// TIA Portal project "proiect" (V17) (continued)
   // ASSB[18] := 18;
   // ASSB[19] := 19;
   // ASSB[20] := 20;
   // ASSB[21] := 21;
   // ASSB[22] := 22;
   // ASSB[23] := 23;
   // ASSB[24] := 24;
   // ASSB[25] := 25;
   // ASSB[26] := 26;
   // ASSB[27] := 27;
   // ASSB[28] := 28;
   // ASSB[29] := 29;
   // ASSB[30] := 30;
   // ASSB[31] := 31;
   // ASSB[32] := 32;
   // ASSB[33] := 33;
   // ASSB[34] := 34;
   // ASSB[35] := 35;
   // ASSB[36] := 36;
   // ASSB[37] := 37;
   // ASSB[38] := 38;
   // ASSB[39] := 39;
   // ASSB[40] := 40;
   // ASSB[41] := 41;
   // ASSB[42] := 42;
   // ASSB[43] := 43;
   // ASSB[44] := 44;
   // ASSB[45] := 45;
   // ASSB[46] := 46;
   // ASSB[47] := 47;
   // ASSB[48] := 48;
   // ASSB[49] := 49;
   // ASSB[50] := 50;
   // ASSB[51] := 51;
   // ASSB[52] := 52;
   // ASSB[53] := 53;
   // ASSB[54] := 54;
   // ASSB[55] := 55;
   // ASSB[56] := 56;
   // ASSB[57] := 57;
   // ASSB[58] := 58;
   // ASSB[59] := 59;
   // ASSB[60] := 60;
   // ASSB[61] := 61;
   // ASSB[62] := 62;
   // ASSB[63] := 63;
   // ASSB[64] := 64;
   // ASSB[65] := 65;
   // ASSB[66] := 66;
   // ASSB[67] := 67;
   // ASSB[68] := 68;
   // ASSB[69] := 69;
   // ASSB[70] := 70;
   // ASSB[71] := 71;
   // ASSB[72] := 72;
   // ASSB[73] := 73;
   // ASSB[74] := 74;
   // ASSB[75] := 75;
   // ASSB[76] := 76;
   // ASSB[77] := 77;
   // PTTS[5] := 2;
   // PTTS[6] := 3;
   // PTTS[7] := 4;
   // PTTS[8] := 5;
   // PTTS[9] := 6;
   // PTTS[10] := 7;
   // PTTS[11] := 72;
   // PTTS[12] := 9;
   // PTTS[13] := 10;
   // PTTS[14] := 11;
   // PTTS[15] := 98;
   // PTTS[16] := 13;
   // PTTS[17] := 14;
   // PTTS[18] := 15;
   // PTTS[19] := 16;
   // PTTS[20] := 17;
   // PTTS[21] := 19;
   // PTTS[22] := 20;
   // PTTS[23] := 21;
   // PTTS[24] := 22;
   // PTTS[25] := 23;
   // PTTS[26] := 24;
   // PTTS[27] := 69;
   // PTTS[28] := 26;
   // PTTS[29] := 27;
   // PTTS[30] := 28;
   // PTTS[31] := 97;
   // PTTS[32] := 30;
   // PTTS[33] := 31;
   // PTTS[34] := 32;
   // PTTS[35] := 33;
   // PTTS[36] := 34;
   // PTTS[37] := 36;
   // PTTS[38] := 37;
   // PTTS[39] := 38;
   // PTTS[40] := 68;
   // PTTS[41] := 40;
   // PTTS[42] := 41;
   // PTTS[43] := 42;
   // PTTS[44] := 96;
   // PTTS[45] := 44;
   // PTTS[46] := 45;
   // PTTS[47] := 46;
   // PTTS[48] := 47;
   // PTTS[49] := 48;
   // PTTS[50] := 53;
   // PTTS[51] := 55;
   // PTTS[52] := 99;
   // PTTS[53] := 57;
   // PTTS[54] := 58;
   // PTTS[55] := 54;
   // PTTS[56] := 59;
   // PTTS[57] := 60;
   // PTTS[58] := 255;
   // PTTS[59] := 62;
   // PTTS[60] := 39;
   // PTTS[61] := 64;
   // PTTS[62] := 66;
   // PTTS[63] := 67;
   // PTTS[64] := 8;
   // PTTS[65] := 25;
   // PTTS[66] := 70;
   // PTTS[67] := 71;
   // PTTS[68] := 73;
   // PTTS[69] := 74;
   // PTTS[70] := 1;
   // PTTS[71] := 63;
   // PTTS[72] := 76;
   // PTTS[73] := 78;
   // PTTS[74] := 43;
   // PTTS[75] := 49;
   // PTTS[76] := 80;
   // PTTS[77] := 29;
   // NTTS[5] := 3;
   // NTTS[6] := 4;
   // NTTS[7] := 5;
   // NTTS[8] := 6;
   // NTTS[9] := 7;
   // NTTS[10] := 8;
   // NTTS[11] := 9;
   // NTTS[12] := 10;
   // NTTS[13] := 11;
   // NTTS[14] := 12;
   // NTTS[15] := 13;
   // NTTS[16] := 14;
   // NTTS[17] := 15;
   // NTTS[18] := 16;
   // NTTS[19] := 17;
   // NTTS[20] := 18;
   // NTTS[21] := 20;
   // NTTS[22] := 21;
   // NTTS[23] := 22;
   // NTTS[24] := 23;
   // NTTS[25] := 24;
   // NTTS[26] := 25;
   // NTTS[27] := 26;
   // NTTS[28] := 27;
   // NTTS[29] := 28;
   // NTTS[30] := 29;
   // NTTS[31] := 30;
   // NTTS[32] := 31;
   // NTTS[33] := 32;
   // NTTS[34] := 33;
   // NTTS[35] := 34;
   // NTTS[36] := 35;
   // NTTS[37] := 37;
   // NTTS[38] := 38;
   // NTTS[39] := 39;
   // NTTS[40] := 40;
   // NTTS[41] := 41;
   // NTTS[42] := 42;
   // NTTS[43] := 78;
   // NTTS[44] := 44;
   // NTTS[45] := 45;
   // NTTS[46] := 46;
   // NTTS[47] := 47;
   // NTTS[48] := 48;
   // NTTS[49] := 49;
   // NTTS[50] := 55;
   // NTTS[51] := 56;
   // NTTS[52] := 57;
   // NTTS[53] := 58;
   // NTTS[54] := 54;
   // NTTS[55] := 59;
   // NTTS[56] := 60;
   // NTTS[57] := 61;
   // NTTS[58] := 62;
   // NTTS[59] := 63;
   // NTTS[60] := 66;
   // NTTS[61] := 65;
   // NTTS[62] := 67;
   // NTTS[63] := 68;
   // NTTS[64] := 73;
   // NTTS[65] := 70;
   // NTTS[66] := 71;
   // NTTS[67] := 69;
   // NTTS[68] := 74;
   // NTTS[69] := 72;
   // NTTS[70] := 36;
   // NTTS[71] := 76;
   // NTTS[72] := 77;
   // NTTS[73] := 43;
   // NTTS[74] := 79;
   // NTTS[75] := 80;
   // NTTS[76] := 81;
   // NTTS[77] := 82;
   // SW_SQTS[3] := 2;
   // SW_SQTS[4] := 2;
   // SW_SQTS[5] := 3;
   // SW_SQTS[6] := 3;
   // SW_SQTS[7] := 3;
   // SW_SQTS[8] := 3;
   // SW_SQTS[9] := 3;
   // SW_SQTS[10] := 3;
   // SW_SQTS[11] := 3;
   // SW_SQTS[12] := 3;
   // SW_SQTS[13] := 3;
   // SW_SQTS[14] := 3;
   // SW_SQTS[15] := 3;
   // SW_SQTS[16] := 3;
   // SW_SQTS[17] := 3;
   // SW_SQTS[18] := 3;
   // SW_SQTS[19] := 3;
   // SW_SQTS[20] := 3;
   // SW_SQTS[21] := 4;
   // SW_SQTS[22] := 4;
   // SW_SQTS[23] := 4;
   // SW_SQTS[24] := 4;
   // SW_SQTS[25] := 4;
   // SW_SQTS[26] := 4;
   // SW_SQTS[27] := 4;
   // SW_SQTS[28] := 4;
   // SW_SQTS[29] := 4;
   // SW_SQTS[30] := 4;
   // SW_SQTS[31] := 4;
   // SW_SQTS[32] := 4;
   // SW_SQTS[33] := 4;
   // SW_SQTS[34] := 4;
   // SW_SQTS[35] := 4;
   // SW_SQTS[36] := 4;
   // SW_SQTS[37] := 5;
   // SW_SQTS[38] := 5;
   // SW_SQTS[39] := 5;
   // SW_SQTS[40] := 5;
   // SW_SQTS[41] := 5;
   // SW_SQTS[42] := 5;
   // SW_SQTS[43] := 5;
   // SW_SQTS[44] := 5;
   // SW_SQTS[45] := 5;
   // SW_SQTS[46] := 5;
   // SW_SQTS[47] := 5;
   // SW_SQTS[48] := 5;
   // SW_SQTS[49] := 5;
   // SW_SQTS[50] := 2;
   // SW_SQTS[51] := 2;
   // SW_SQTS[52] := 2;
   // SW_SQTS[53] := 2;
   // SW_SQTS[54] := 2;
   // SW_SQTS[55] := 2;
   // SW_SQTS[56] := 2;
   // SW_SQTS[57] := 2;
   // SW_SQTS[58] := 6;
   // SW_SQTS[59] := 7;
   // SW_SQTS[60] := 5;
   // SW_SQTS[61] := 8;
   // SW_SQTS[62] := 5;
   // SW_SQTS[63] := 5;
   // SW_SQTS[64] := 3;
   // SW_SQTS[65] := 4;
   // SW_SQTS[66] := 4;
   // SW_SQTS[67] := 4;
   // SW_SQTS[68] := 3;
   // SW_SQTS[69] := 3;
   // SW_SQTS[70] := 9;
   // SW_SQTS[71] := 7;
   // SW_SQTS[72] := 7;
   // SW_SQTS[73] := 5;
   // SW_SQTS[74] := 5;
   // SW_SQTS[75] := 5;
   // SW_SQTS[76] := 5;
   // SW_SQTS[77] := 4;
   // SINI[2] := 255;
   // LSTT[83] := 255;
   // LSTT[84] := 255;
   // LSTT[86] := 255;
   // ATAJ[82] := 82;
   // ATAJ[83] := 83;
   // ATAJ[84] := 84;
   // ATAJ[85] := 85;
   // ATAJ[86] := 86;
   // ATAB[82] := 82;
   // ATAB[83] := 83;
   // ATAB[84] := 84;
   // ATAB[85] := 85;
   // ATAB[86] := 86;
   // PSTT[82] := 77;
   // PSTT[83] := 78;
   // PSTT[84] := 79;
   // PSTT[85] := 80;
   // PSTT[86] := 81;
   // NSTT[83] := 91;
   // NSTT[84] := 80;
   // NSTT[86] := 82;
   // ASSJ[78] := 78;
   // ASSJ[79] := 79;
   // ASSJ[80] := 80;
   // ASSJ[81] := 81;
   // ASSB[78] := 78;
   // ASSB[79] := 79;
   // ASSB[80] := 80;
   // ASSB[81] := 81;
   // PTTS[78] := 82;
   // PTTS[79] := 35;
   // PTTS[80] := 84;
   // PTTS[81] := 12;
   // NTTS[78] := 83;
   // NTTS[79] := 84;
   // NTTS[80] := 85;
   // NTTS[81] := 86;
   // SW_SQTS[78] := 4;
   // SW_SQTS[79] := 4;
   // SW_SQTS[80] := 4;
   // SW_SQTS[81] := 3;
   // SWITCH[0] := 192;
   // SWITCH[1] := 1;
   // SWITCH[2] := 14;
   // SWITCH[3] := 112;
   // SWITCH[4] := 128;
   // SWITCH[5] := 3;
   // SWITCH[6] := 28;
   // SWITCH[7] := 224;
   // LSTT[87] := 255;
   // LSTT[88] := 255;
   // LSTT[90] := 255;
   // LSTT[91] := 255;
   // LSTT[92] := 255;
   // LSTT[94] := 255;
   // ATAJ[87] := 87;
   // ATAJ[88] := 88;
   // ATAJ[89] := 89;
   // ATAJ[90] := 90;
   // ATAJ[91] := 91;
   // ATAJ[92] := 92;
   // ATAJ[93] := 93;
   // ATAJ[94] := 94;
   // ATAJ[95] := 95;
   // ATAB[87] := 87;
   // ATAB[88] := 88;
   // ATAB[89] := 89;
   // ATAB[90] := 90;
   // ATAB[91] := 91;
   // ATAB[92] := 92;
   // ATAB[93] := 93;
   // ATAB[95] := 95;
   // PSTT[87] := 82;
   // PSTT[88] := 83;
   // PSTT[89] := 84;
   // PSTT[90] := 85;
   // PSTT[91] := 86;
   // PSTT[92] := 87;
   // PSTT[93] := 88;
   // PSTT[95] := 89;
   // NSTT[87] := 92;
   // NSTT[88] := 84;
   // NSTT[90] := 86;
   // NSTT[91] := 93;
   // NSTT[92] := 88;
   // NSTT[94] := 89;
   // ASSJ[82] := 82;
   // ASSJ[83] := 83;
   // ASSJ[84] := 84;
   // ASSJ[85] := 85;
   // ASSJ[86] := 86;
   // ASSJ[87] := 87;
   // ASSJ[88] := 88;
   // ASSJ[89] := 89;
   // ASSB[82] := 82;
   // ASSB[83] := 83;
   // ASSB[84] := 84;
   // ASSB[85] := 85;
   // ASSB[86] := 86;
   // ASSB[87] := 87;
   // ASSB[88] := 88;
   // ASSB[89] := 89;
   // PTTS[82] := 86;
   // PTTS[83] := 18;
   // PTTS[84] := 88;
   // PTTS[85] := 56;
   // PTTS[86] := 90;
   // PTTS[87] := 61;
   // PTTS[88] := 92;
   // PTTS[89] := 94;
   // NTTS[82] := 87;
   // NTTS[83] := 88;
   // NTTS[84] := 89;
   // NTTS[85] := 90;
   // NTTS[86] := 91;
   // NTTS[87] := 92;
   // NTTS[88] := 93;
   // NTTS[89] := 95;
   // SW_SQTS[82] := 3;
   // SW_SQTS[83] := 3;
   // SW_SQTS[84] := 3;
   // SW_SQTS[85] := 2;
   // SW_SQTS[86] := 2;
   // SW_SQTS[87] := 2;
   // SW_SQTS[88] := 2;
   // SW_SQTS[89] := 10;
   // SW_SQTS[2] := 2;
   // SWITCH[8] := 252;
   // SWITCH[9] := 248;
   // SWITCH[10] := 199;
   // SW_SQTS[1] := 1;
   // ATAB[0] := 94;
   // SWITCH[12] := 6;
   // LSTT[61] := 255;
   // LSTT[43] := 255;
   // LSTT[22] := 255;
   // SWITCH[11] := 63;
   // NSTT[61] := 87;
   // NSTT[43] := 74;
   // NSTT[22] := 24;
   // SWITCH[13] := 14;
   // SWITCH[14] := 112;
   // LSTT[96] := 255;
   // LSTT[97] := 255;
   // LSTT[98] := 255;
   // LSTT[99] := 255;
   // ATAJ[96] := 96;
   // ATAJ[97] := 97;
   // ATAJ[98] := 98;
   // ATAJ[99] := 99;
   // ATAB[96] := 96;
   // ATAB[97] := 97;
   // ATAB[98] := 98;
   // ATAB[99] := 99;
   // PSTT[96] := 90;
   // PSTT[97] := 91;
   // PSTT[98] := 92;
   // PSTT[99] := 93;
   // NSTT[96] := 44;
   // NSTT[97] := 31;
   // NSTT[98] := 15;
   // NSTT[99] := 52;
   // ASSJ[90] := 90;
   // ASSJ[91] := 91;
   // ASSJ[92] := 92;
   // ASSJ[93] := 93;
   // ASSB[90] := 90;
   // ASSB[91] := 91;
   // ASSB[92] := 92;
   // ASSB[93] := 93;
   // PTTS[90] := 79;
   // PTTS[91] := 83;
   // PTTS[92] := 87;
   // PTTS[93] := 91;
   // NTTS[90] := 96;
   // NTTS[91] := 97;
   // NTTS[92] := 98;
   // NTTS[93] := 99;
   // SW_SQTS[90] := 5;
   // SW_SQTS[91] := 4;
   // SW_SQTS[92] := 3;
   // SW_SQTS[93] := 2;
BEGIN
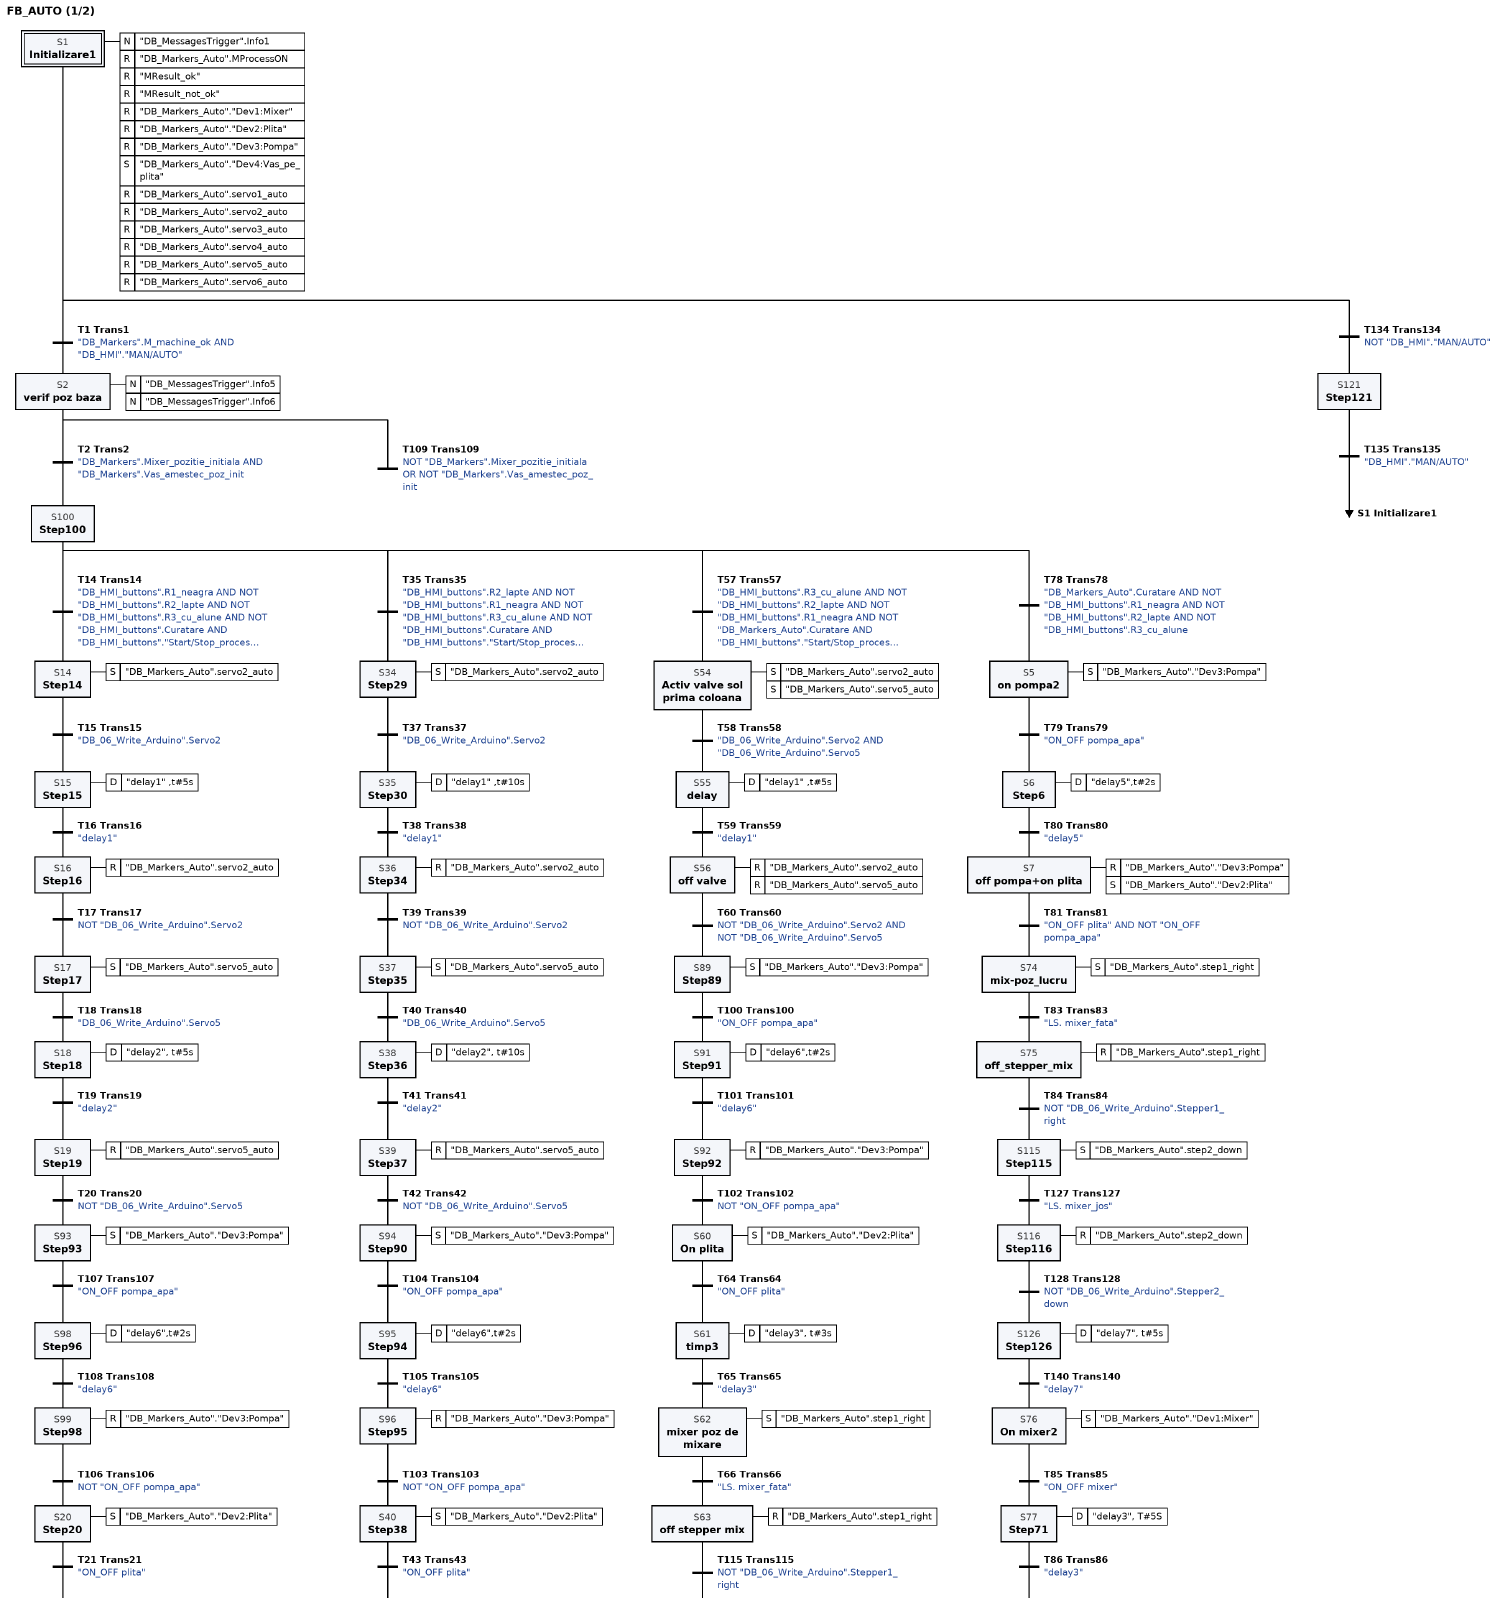
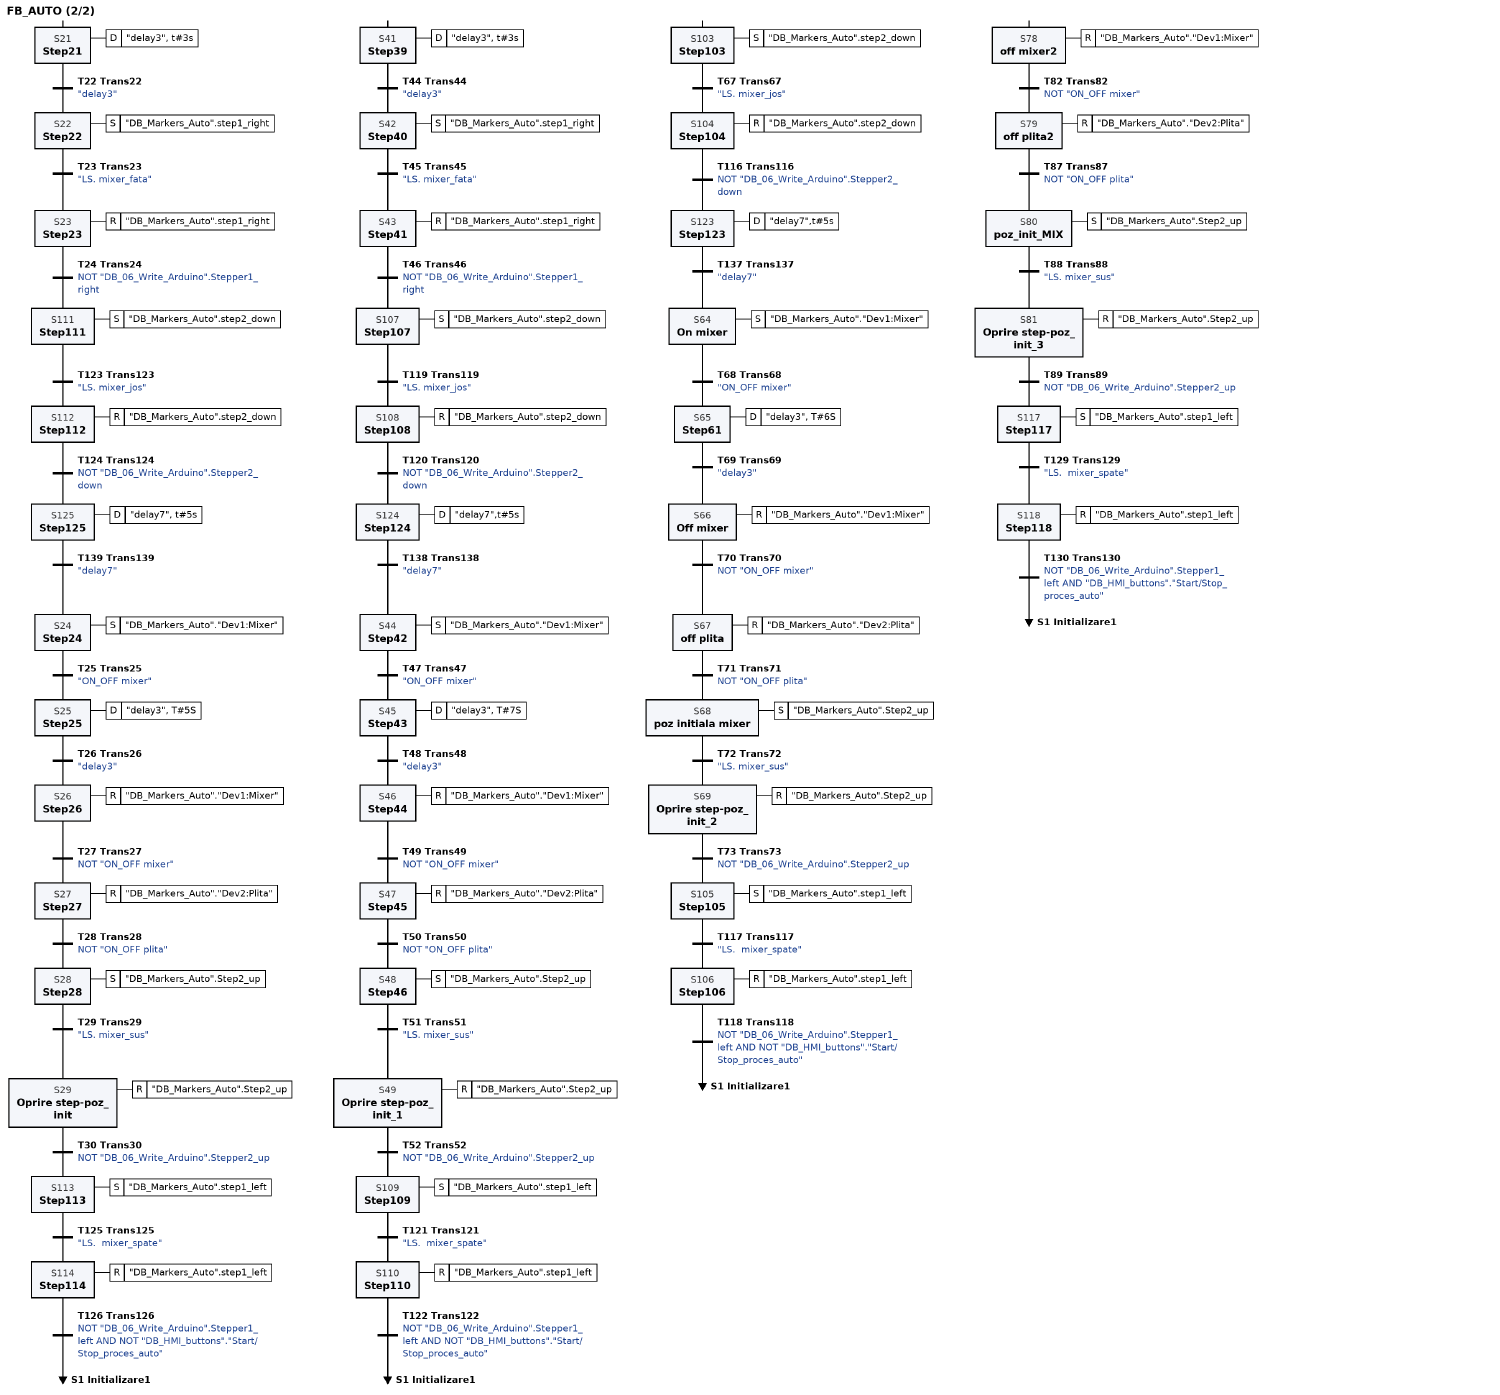
   // sequencer 1
   INITIAL_STEP Initializare1:   // S1, max time T#10S, warning time T#7S
      // Initializare
              N    "DB_MessagesTrigger".Info1
              R    "DB_Markers_Auto".MProcessON
              R    "MResult_ok"
              R    "MResult_not_ok"
              R    "DB_Markers_Auto"."Dev1:Mixer"
              R    "DB_Markers_Auto"."Dev2:Plita"
              R    "DB_Markers_Auto"."Dev3:Pompa"
              S    "DB_Markers_Auto"."Dev4:Vas_pe_plita"
              R    "DB_Markers_Auto".servo1_auto
              R    "DB_Markers_Auto".servo2_auto
              R    "DB_Markers_Auto".servo3_auto
              R    "DB_Markers_Auto".servo4_auto
              R    "DB_Markers_Auto".servo5_auto
              R    "DB_Markers_Auto".servo6_auto
              R    "DB_Markers_Auto".step1_left
              R    "DB_Markers_Auto".step1_right
              R    "DB_Markers_Auto".Step2_up
              R    "DB_Markers_Auto".step2_down
   END_STEP
   TRANSITION Trans1 FROM Initializare1 TO "verif poz baza"   // T1
      := "DB_Markers".M_machine_ok AND "DB_HMI"."MAN/AUTO";
   END_TRANSITION
   TRANSITION Trans134 FROM Initializare1 TO Step121   // T134
      := NOT "DB_HMI"."MAN/AUTO";
   END_TRANSITION
   STEP "verif poz baza":   // S2, max time T#10S, warning time T#7S
      // Verificare dispozitive in pozitia de baza
              N    "DB_MessagesTrigger".Info5
              N    "DB_MessagesTrigger".Info6
   END_STEP
   TRANSITION Trans2 FROM "verif poz baza" TO Step100   // T2
      := "DB_Markers".Mixer_pozitie_initiala AND "DB_Markers".Vas_amestec_poz_init;
   END_TRANSITION
   TRANSITION Trans109 FROM "verif poz baza" TO ?   // T109
      := NOT "DB_Markers".Mixer_pozitie_initiala OR NOT "DB_Markers".Vas_amestec_poz_init;
   END_TRANSITION
   STEP Step103:   // S103, max time T#10S, warning time T#7S
              S    "DB_Markers_Auto".step2_down
   END_STEP
   TRANSITION Trans67 FROM Step103 TO Step104   // T67
      := "LS. mixer_jos";
   END_TRANSITION
   STEP Step29:   // S34, max time T#10S, warning time T#7S
      // Activare valve solutii rand superior
              S    "DB_Markers_Auto".servo2_auto
   END_STEP
   TRANSITION Trans37 FROM Step29 TO Step30   // T37
      := "DB_06_Write_Arduino".Servo2;
   END_TRANSITION
   STEP Step14:   // S14, max time T#10S, warning time T#7S
      // Activare valve solutii rand superior
              S    "DB_Markers_Auto".servo2_auto
   END_STEP
   TRANSITION Trans15 FROM Step14 TO Step15   // T15
      := "DB_06_Write_Arduino".Servo2;
   END_TRANSITION
   STEP Step15:   // S15, max time T#10S, warning time T#7S
      // delay
              D    "delay1" ,t#5s
   END_STEP
   TRANSITION Trans16 FROM Step15 TO Step16   // T16
      := "delay1";
   END_TRANSITION
   STEP Step16:   // S16, max time T#10S, warning time T#7S
      // inchidere valve rand superior
              R    "DB_Markers_Auto".servo2_auto
   END_STEP
   TRANSITION Trans17 FROM Step16 TO Step17   // T17
      := NOT "DB_06_Write_Arduino".Servo2;
   END_TRANSITION
   STEP Step17:   // S17, max time T#10S, warning time T#7S
      // deschidere valve solutii rand inferior
              S    "DB_Markers_Auto".servo5_auto
   END_STEP
   TRANSITION Trans18 FROM Step17 TO Step18   // T18
      := "DB_06_Write_Arduino".Servo5;
   END_TRANSITION
   STEP Step18:   // S18, max time T#10S, warning time T#7S
      // delay
              D    "delay2", t#5s
   END_STEP
   TRANSITION Trans19 FROM Step18 TO Step19   // T19
      := "delay2";
   END_TRANSITION
   STEP Step19:   // S19, max time T#10S, warning time T#7S
      // inchidere valve rand inferior
              R    "DB_Markers_Auto".servo5_auto
   END_STEP
   TRANSITION Trans20 FROM Step19 TO Step93   // T20
      := NOT "DB_06_Write_Arduino".Servo5;
   END_TRANSITION
   STEP Step20:   // S20, max time T#10S, warning time T#7S
      // deschidere plita
              S    "DB_Markers_Auto"."Dev2:Plita"
   END_STEP
   TRANSITION Trans21 FROM Step20 TO Step21   // T21
      := "ON_OFF plita";
   END_TRANSITION
   STEP Step21:   // S21, max time T#10S, warning time T#7S
      // delay
              D    "delay3", t#3s
   END_STEP
   TRANSITION Trans22 FROM Step21 TO Step22   // T22
      := "delay3";
   END_TRANSITION
   STEP Step22:   // S22, max time T#10S, warning time T#7S
      // pozitionare mixer/pornire stepper
              S    "DB_Markers_Auto".step1_right
   END_STEP
   TRANSITION Trans23 FROM Step22 TO Step23   // T23
      := "LS. mixer_fata";
   END_TRANSITION
   STEP Step23:   // S23, max time T#10S, warning time T#7S
      // Oprire stepper/mixer
              R    "DB_Markers_Auto".step1_right
   END_STEP
   TRANSITION Trans24 FROM Step23 TO Step111   // T24
      := NOT "DB_06_Write_Arduino".Stepper1_right;
   END_TRANSITION
   STEP Step24:   // S24, max time T#10S, warning time T#7S
      // Pornire mixer(on,off)
              S    "DB_Markers_Auto"."Dev1:Mixer"
   END_STEP
   TRANSITION Trans25 FROM Step24 TO Step25   // T25
      := "ON_OFF mixer";
   END_TRANSITION
   STEP Step25:   // S25, max time T#10S, warning time T#7S
      // Delay(timp de mixare)
              D    "delay3", T#5S
   END_STEP
   TRANSITION Trans26 FROM Step25 TO Step26   // T26
      := "delay3";
   END_TRANSITION
   STEP Step26:   // S26, max time T#10S, warning time T#7S
      // Oprire mixer
              R    "DB_Markers_Auto"."Dev1:Mixer"
   END_STEP
   TRANSITION Trans27 FROM Step26 TO Step27   // T27
      := NOT "ON_OFF mixer";
   END_TRANSITION
   STEP Step27:   // S27, max time T#10S, warning time T#7S
      // Oprire plita
              R    "DB_Markers_Auto"."Dev2:Plita"
   END_STEP
   TRANSITION Trans28 FROM Step27 TO Step28   // T28
      := NOT "ON_OFF plita";
   END_TRANSITION
   STEP Step28:   // S28, max time T#10S, warning time T#7S
      // RETRAGERE MIXER IN POZITIA INITIALA
              S    "DB_Markers_Auto".Step2_up
   END_STEP
   TRANSITION Trans29 FROM Step28 TO "Oprire step-poz_init"   // T29
      := "LS. mixer_sus";
   END_TRANSITION
   STEP "Oprire step-poz_init":   // S29, max time T#10S, warning time T#7S
      // Oprire Stepper_pozitie initiala
              R    "DB_Markers_Auto".Step2_up
   END_STEP
   TRANSITION Trans30 FROM "Oprire step-poz_init" TO Step113   // T30
      := NOT "DB_06_Write_Arduino".Stepper2_up;
   END_TRANSITION
   STEP Step30:   // S35, max time T#10S, warning time T#7S
      // delay
              D    "delay1" ,t#10s
   END_STEP
   TRANSITION Trans38 FROM Step30 TO Step34   // T38
      := "delay1";
   END_TRANSITION
   STEP Step34:   // S36, max time T#10S, warning time T#7S
      // inchidere valve rand superior
              R    "DB_Markers_Auto".servo2_auto
   END_STEP
   TRANSITION Trans39 FROM Step34 TO Step35   // T39
      := NOT "DB_06_Write_Arduino".Servo2;
   END_TRANSITION
   STEP Step35:   // S37, max time T#10S, warning time T#7S
      // deschidere valve solutii rand inferior
              S    "DB_Markers_Auto".servo5_auto
   END_STEP
   TRANSITION Trans40 FROM Step35 TO Step36   // T40
      := "DB_06_Write_Arduino".Servo5;
   END_TRANSITION
   STEP Step36:   // S38, max time T#10S, warning time T#7S
      // delay
              D    "delay2", t#10s
   END_STEP
   TRANSITION Trans41 FROM Step36 TO Step37   // T41
      := "delay2";
   END_TRANSITION
   STEP Step37:   // S39, max time T#10S, warning time T#7S
      // inchidere valve rand inferior
              R    "DB_Markers_Auto".servo5_auto
   END_STEP
   TRANSITION Trans42 FROM Step37 TO Step90   // T42
      := NOT "DB_06_Write_Arduino".Servo5;
   END_TRANSITION
   STEP Step38:   // S40, max time T#10S, warning time T#7S
      // deschidere plita
              S    "DB_Markers_Auto"."Dev2:Plita"
   END_STEP
   TRANSITION Trans43 FROM Step38 TO Step39   // T43
      := "ON_OFF plita";
   END_TRANSITION
   STEP Step39:   // S41, max time T#10S, warning time T#7S
      // delay
              D    "delay3", t#3s
   END_STEP
   TRANSITION Trans44 FROM Step39 TO Step40   // T44
      := "delay3";
   END_TRANSITION
   STEP Step40:   // S42, max time T#10S, warning time T#7S
      // pozitionare mixer/pornire stepper
              S    "DB_Markers_Auto".step1_right
   END_STEP
   TRANSITION Trans45 FROM Step40 TO Step41   // T45
      := "LS. mixer_fata";
   END_TRANSITION
   STEP Step41:   // S43, max time T#10S, warning time T#7S
      // Oprire stepper/mixer
              R    "DB_Markers_Auto".step1_right
   END_STEP
   TRANSITION Trans46 FROM Step41 TO Step107   // T46
      := NOT "DB_06_Write_Arduino".Stepper1_right;
   END_TRANSITION
   STEP Step42:   // S44, max time T#10S, warning time T#7S
      // Pornire mixer(on,off)
              S    "DB_Markers_Auto"."Dev1:Mixer"
   END_STEP
   TRANSITION Trans47 FROM Step42 TO Step43   // T47
      := "ON_OFF mixer";
   END_TRANSITION
   STEP Step43:   // S45, max time T#10S, warning time T#7S
      // Delay(timp de mixare)
              D    "delay3", T#7S
   END_STEP
   TRANSITION Trans48 FROM Step43 TO Step44   // T48
      := "delay3";
   END_TRANSITION
   STEP Step44:   // S46, max time T#10S, warning time T#7S
      // Oprire mixer
              R    "DB_Markers_Auto"."Dev1:Mixer"
   END_STEP
   TRANSITION Trans49 FROM Step44 TO Step45   // T49
      := NOT "ON_OFF mixer";
   END_TRANSITION
   STEP Step45:   // S47, max time T#10S, warning time T#7S
      // Oprire plita
              R    "DB_Markers_Auto"."Dev2:Plita"
   END_STEP
   TRANSITION Trans50 FROM Step45 TO Step46   // T50
      := NOT "ON_OFF plita";
   END_TRANSITION
   STEP Step46:   // S48, max time T#10S, warning time T#7S
      // RETRAGERE MIXER IN POZITIA INITIALA
              S    "DB_Markers_Auto".Step2_up
   END_STEP
   TRANSITION Trans51 FROM Step46 TO "Oprire step-poz_init_1"   // T51
      := "LS. mixer_sus";
   END_TRANSITION
   STEP "Oprire step-poz_init_1":   // S49, max time T#10S, warning time T#7S
      // Oprire Stepper_pozitie initiala
              R    "DB_Markers_Auto".Step2_up
   END_STEP
   TRANSITION Trans52 FROM "Oprire step-poz_init_1" TO Step109   // T52
      := NOT "DB_06_Write_Arduino".Stepper2_up;
   END_TRANSITION
   STEP "Activ valve sol prima coloana":   // S54, max time T#10S, warning time T#7S
      // Activare valve solutii prima coloana
              S    "DB_Markers_Auto".servo2_auto
              S    "DB_Markers_Auto".servo5_auto
   END_STEP
   TRANSITION Trans58 FROM "Activ valve sol prima coloana" TO delay   // T58
      := "DB_06_Write_Arduino".Servo2 AND "DB_06_Write_Arduino".Servo5;
   END_TRANSITION
   STEP delay:   // S55, max time T#10S, warning time T#7S
      // delay
              D    "delay1" ,t#5s
   END_STEP
   TRANSITION Trans59 FROM delay TO "off valve"   // T59
      := "delay1";
   END_TRANSITION
   STEP "off valve":   // S56, max time T#10S, warning time T#7S
      // inchidere valve coloana 1
              R    "DB_Markers_Auto".servo2_auto
              R    "DB_Markers_Auto".servo5_auto
   END_STEP
   TRANSITION Trans60 FROM "off valve" TO Step89   // T60
      := NOT "DB_06_Write_Arduino".Servo2 AND NOT "DB_06_Write_Arduino".Servo5;
   END_TRANSITION
   STEP "On plita":   // S60, max time T#10S, warning time T#7S
      // deschidere plita
              S    "DB_Markers_Auto"."Dev2:Plita"
   END_STEP
   TRANSITION Trans64 FROM "On plita" TO timp3   // T64
      := "ON_OFF plita";
   END_TRANSITION
   STEP timp3:   // S61, max time T#10S, warning time T#7S
      // delay
              D    "delay3", t#3s
   END_STEP
   TRANSITION Trans65 FROM timp3 TO "mixer poz de mixare"   // T65
      := "delay3";
   END_TRANSITION
   STEP "mixer poz de mixare":   // S62, max time T#10S, warning time T#7S
      // pozitionare mixer/pornire stepper
              S    "DB_Markers_Auto".step1_right
   END_STEP
   TRANSITION Trans66 FROM "mixer poz de mixare" TO "off stepper mix"   // T66
      := "LS. mixer_fata";
   END_TRANSITION
   STEP "off stepper mix":   // S63, max time T#10S, warning time T#7S
      // Oprire stepper/mixer
              R    "DB_Markers_Auto".step1_right
   END_STEP
   TRANSITION Trans115 FROM "off stepper mix" TO Step103   // T115
      := NOT "DB_06_Write_Arduino".Stepper1_right;
   END_TRANSITION
   STEP "On mixer":   // S64, max time T#10S, warning time T#7S
      // Pornire mixer(on,off)
              S    "DB_Markers_Auto"."Dev1:Mixer"
   END_STEP
   TRANSITION Trans68 FROM "On mixer" TO Step61   // T68
      := "ON_OFF mixer";
   END_TRANSITION
   STEP Step61:   // S65, max time T#10S, warning time T#7S
      // Delay(timp de mixare)
              D    "delay3", T#6S
   END_STEP
   TRANSITION Trans69 FROM Step61 TO "Off mixer"   // T69
      := "delay3";
   END_TRANSITION
   STEP "Off mixer":   // S66, max time T#10S, warning time T#7S
      // Oprire mixer
              R    "DB_Markers_Auto"."Dev1:Mixer"
   END_STEP
   TRANSITION Trans70 FROM "Off mixer" TO "off plita"   // T70
      := NOT "ON_OFF mixer";
   END_TRANSITION
   STEP "off plita":   // S67, max time T#10S, warning time T#7S
      // Oprire plita
              R    "DB_Markers_Auto"."Dev2:Plita"
   END_STEP
   TRANSITION Trans71 FROM "off plita" TO "poz initiala mixer"   // T71
      := NOT "ON_OFF plita";
   END_TRANSITION
   STEP "poz initiala mixer":   // S68, max time T#10S, warning time T#7S
      // RETRAGERE MIXER IN POZITIA INITIALA
              S    "DB_Markers_Auto".Step2_up
   END_STEP
   TRANSITION Trans72 FROM "poz initiala mixer" TO "Oprire step-poz_init_2"   // T72
      := "LS. mixer_sus";
   END_TRANSITION
   STEP "Oprire step-poz_init_2":   // S69, max time T#10S, warning time T#7S
      // Oprire Stepper_pozitie initiala
              R    "DB_Markers_Auto".Step2_up
   END_STEP
   TRANSITION Trans73 FROM "Oprire step-poz_init_2" TO Step105   // T73
      := NOT "DB_06_Write_Arduino".Stepper2_up;
   END_TRANSITION
   STEP "on pompa2":   // S5, max time T#10S, warning time T#7S
      // curatare(activare pompa+incalzire plita+mixare)
              S    "DB_Markers_Auto"."Dev3:Pompa"
   END_STEP
   TRANSITION Trans79 FROM "on pompa2" TO Step6   // T79
      := "ON_OFF pompa_apa";
   END_TRANSITION
   STEP Step6:   // S6, max time T#10S, warning time T#7S
      // delay
              D    "delay5",t#2s
   END_STEP
   TRANSITION Trans80 FROM Step6 TO "off pompa+on plita"   // T80
      := "delay5";
   END_TRANSITION
   STEP "off pompa+on plita":   // S7, max time T#10S, warning time T#7S
      // oprire pompa+activare plita
              R    "DB_Markers_Auto"."Dev3:Pompa"
              S    "DB_Markers_Auto"."Dev2:Plita"
   END_STEP
   TRANSITION Trans81 FROM "off pompa+on plita" TO "mix-poz_lucru"   // T81
      := "ON_OFF plita" AND NOT "ON_OFF pompa_apa";
   END_TRANSITION
   STEP "Oprire step-poz_init_3":   // S81, max time T#10S, warning time T#7S
      // Oprire Stepper_pozitie initiala
              R    "DB_Markers_Auto".Step2_up
   END_STEP
   TRANSITION Trans89 FROM "Oprire step-poz_init_3" TO Step117   // T89
      := NOT "DB_06_Write_Arduino".Stepper2_up;
   END_TRANSITION
   STEP "mix-poz_lucru":   // S74, max time T#10S, warning time T#7S
      // pozitionare mixer/pornire stepper
              S    "DB_Markers_Auto".step1_right
   END_STEP
   TRANSITION Trans83 FROM "mix-poz_lucru" TO off_stepper_mix   // T83
      := "LS. mixer_fata";
   END_TRANSITION
   STEP off_stepper_mix:   // S75, max time T#10S, warning time T#7S
      // Oprire stepper/mixer
              R    "DB_Markers_Auto".step1_right
   END_STEP
   TRANSITION Trans84 FROM off_stepper_mix TO Step115   // T84
      := NOT "DB_06_Write_Arduino".Stepper1_right;
   END_TRANSITION
   STEP "On mixer2":   // S76, max time T#10S, warning time T#7S
      // Pornire mixer(on,off)
              S    "DB_Markers_Auto"."Dev1:Mixer"
   END_STEP
   TRANSITION Trans85 FROM "On mixer2" TO Step71   // T85
      := "ON_OFF mixer";
   END_TRANSITION
   STEP Step71:   // S77, max time T#10S, warning time T#7S
      // Delay(timp de mixare)
              D    "delay3", T#5S
   END_STEP
   TRANSITION Trans86 FROM Step71 TO "off mixer2"   // T86
      := "delay3";
   END_TRANSITION
   STEP "off mixer2":   // S78, max time T#10S, warning time T#7S
      // Oprire mixer
              R    "DB_Markers_Auto"."Dev1:Mixer"
   END_STEP
   TRANSITION Trans82 FROM "off mixer2" TO "off plita2"   // T82
      := NOT "ON_OFF mixer";
   END_TRANSITION
   STEP "off plita2":   // S79, max time T#10S, warning time T#7S
      // Oprire plita
              R    "DB_Markers_Auto"."Dev2:Plita"
   END_STEP
   TRANSITION Trans87 FROM "off plita2" TO poz_init_MIX   // T87
      := NOT "ON_OFF plita";
   END_TRANSITION
   STEP poz_init_MIX:   // S80, max time T#10S, warning time T#7S
      // RETRAGERE MIXER IN POZITIA INITIALA
              S    "DB_Markers_Auto".Step2_up
   END_STEP
   TRANSITION Trans88 FROM poz_init_MIX TO "Oprire step-poz_init_3"   // T88
      := "LS. mixer_sus";
   END_TRANSITION
   STEP Step89:   // S89, max time T#10S, warning time T#7S
              S    "DB_Markers_Auto"."Dev3:Pompa"
   END_STEP
   TRANSITION Trans100 FROM Step89 TO Step91   // T100
      := "ON_OFF pompa_apa";
   END_TRANSITION
   STEP Step91:   // S91, max time T#10S, warning time T#7S
              D    "delay6",t#2s
   END_STEP
   TRANSITION Trans101 FROM Step91 TO Step92   // T101
      := "delay6";
   END_TRANSITION
   STEP Step92:   // S92, max time T#10S, warning time T#7S
      // R
              R    "DB_Markers_Auto"."Dev3:Pompa"
   END_STEP
   TRANSITION Trans102 FROM Step92 TO "On plita"   // T102
      := NOT "ON_OFF pompa_apa";
   END_TRANSITION
   STEP Step90:   // S94, max time T#10S, warning time T#7S
              S    "DB_Markers_Auto"."Dev3:Pompa"
   END_STEP
   TRANSITION Trans104 FROM Step90 TO Step94   // T104
      := "ON_OFF pompa_apa";
   END_TRANSITION
   STEP Step94:   // S95, max time T#10S, warning time T#7S
              D    "delay6",t#2s
   END_STEP
   TRANSITION Trans105 FROM Step94 TO Step95   // T105
      := "delay6";
   END_TRANSITION
   STEP Step95:   // S96, max time T#10S, warning time T#7S
      // R
              R    "DB_Markers_Auto"."Dev3:Pompa"
   END_STEP
   TRANSITION Trans103 FROM Step95 TO Step38   // T103
      := NOT "ON_OFF pompa_apa";
   END_TRANSITION
   STEP Step93:   // S93, max time T#10S, warning time T#7S
              S    "DB_Markers_Auto"."Dev3:Pompa"
   END_STEP
   TRANSITION Trans107 FROM Step93 TO Step96   // T107
      := "ON_OFF pompa_apa";
   END_TRANSITION
   STEP Step96:   // S98, max time T#10S, warning time T#7S
              D    "delay6",t#2s
   END_STEP
   TRANSITION Trans108 FROM Step96 TO Step98   // T108
      := "delay6";
   END_TRANSITION
   STEP Step98:   // S99, max time T#10S, warning time T#7S
      // R
              R    "DB_Markers_Auto"."Dev3:Pompa"
   END_STEP
   TRANSITION Trans106 FROM Step98 TO Step20   // T106
      := NOT "ON_OFF pompa_apa";
   END_TRANSITION
   STEP Step100:   // S100, max time T#10S, warning time T#7S
      // selectare reteta
   END_STEP
   TRANSITION Trans14 FROM Step100 TO Step14   // T14: ciocolata neagra
      := "DB_HMI_buttons".R1_neagra AND NOT "DB_HMI_buttons".R2_lapte AND NOT "DB_HMI_buttons".R3_cu_alune AND NOT "DB_HMI_buttons".Curatare AND "DB_HMI_buttons"."Start/Stop_proces_auto";
   END_TRANSITION
   TRANSITION Trans35 FROM Step100 TO Step29   // T35: Ciocolata cu lapte
      := "DB_HMI_buttons".R2_lapte AND NOT "DB_HMI_buttons".R1_neagra AND NOT "DB_HMI_buttons".R3_cu_alune AND NOT "DB_HMI_buttons".Curatare AND "DB_HMI_buttons"."Start/Stop_proces_auto";
   END_TRANSITION
   TRANSITION Trans57 FROM Step100 TO "Activ valve sol prima coloana"   // T57: Ciocolata cu alune
      := "DB_HMI_buttons".R3_cu_alune AND NOT "DB_HMI_buttons".R2_lapte AND NOT "DB_HMI_buttons".R1_neagra AND NOT "DB_Markers_Auto".Curatare AND "DB_HMI_buttons"."Start/Stop_proces_auto";
   END_TRANSITION
   TRANSITION Trans78 FROM Step100 TO "on pompa2"   // T78: Auto curatare
      := "DB_Markers_Auto".Curatare AND NOT "DB_HMI_buttons".R1_neagra AND NOT "DB_HMI_buttons".R2_lapte AND NOT "DB_HMI_buttons".R3_cu_alune;
   END_TRANSITION
   STEP Step104:   // S104, max time T#10S, warning time T#7S
              R    "DB_Markers_Auto".step2_down
   END_STEP
   TRANSITION Trans116 FROM Step104 TO Step123   // T116
      := NOT "DB_06_Write_Arduino".Stepper2_down;
   END_TRANSITION
   STEP Step105:   // S105, max time T#10S, warning time T#7S
              S    "DB_Markers_Auto".step1_left